// TIA Portal project "Blower_Speeds" (V19)
// Project for control of blower speed through variable frequency drive

(* hardware
DEVICE "S7-1200 station_1"  S7-1200 Station
   slot 0: "Rack_0"  S7-1200 Rack  Rack  V1.0
   slot 1: "PLC_1"  CPU 1212C AC/DC/Rly  6ES7 212-1BE40-0XB0  V4.6
DEVICE "HMI_1"  TP1200 Comfort
   slot 0: "HMI_1"  TP1200 Comfort  6AV2 124-0MC01-0AX0  17.0.0.0
   slot 1: "HMI_RT_1"  TP1200 Comfort  6AV2 124-0MC01-0AX0  17.0.0.0
   slot 5: "HMI_1.IE_CP_1"  PROFINET Interface  17.0.0.0
      slot 1: "PROFINET Interface_1"  PROFINET Interface
         slot 1: "Port_1"  Port
         slot 2: "Port_2"  Port
   slot 7: "HMI_1.MPI/DP_CP_1"  MPI/DP Interface  17.0.0.0
*)

// ===== PLC "PLC_1"  CPU 1212C AC/DC/Rly =====

VAR_GLOBAL   // PLC tag table "Inputs"
   "E_Stop" AT %I0.0 : Bool;   // Emergency stop
   "Start" AT %I0.2 : Bool;   // Pushbutton Start NO
   "Increase_Speed" AT %I0.4 : Bool;   // Pushbutton Increase NO
   "Decrease_Speed" AT %I0.3 : Bool;   // Pushbutton Decrease NO
   "Stop" AT %I0.1 : Bool;   // Pushbutton Stop NC
   "Tag_1" AT %M0.0 : Bool;
   "Tag_2" AT %M0.1 : Bool;
END_VAR

VAR_GLOBAL   // PLC tag table "Outputs"
   "Speed_1" AT %Q0.0 : Bool;   // Select Speed 1
   "Speed_2" AT %Q0.1 : Bool;   // Select Speed 2
   "Speed_3" AT %Q0.2 : Bool;   // Select Speed 3
   "Speed_4" AT %Q0.3 : Bool;   // Select Speed 4
END_VAR

// folder: DB

DATA_BLOCK "Data"   // DB1
TITLE = Data for Set Memories
{ S7_Optimized_Access := 'TRUE' }
AUTHOR : Stiven Perez
VERSION : 0.1
// Data for Set Memories
   VAR
      Start_Stop : Bool;   // Set-Reset Start or Stop Process
      P_Inc : Bool;
      N_Dec : Bool;
      QTime_1 : Bool;
      QTime_2 : Bool;
      QTime_3 : Bool;
      QTime_4 : Bool;
      CV_Speed : Int;
      Reset_Counter : Bool;
   END_VAR
BEGIN
END_DATA_BLOCK

DATA_BLOCK "Start_Stop_DB"   // DB2
{ S7_Optimized_Access := 'TRUE' }
VERSION : 0.1
// stored: InstanceOfName Start_Stop
"Start_Stop"
BEGIN
END_DATA_BLOCK

DATA_BLOCK "Inc_Dec_Speed_DB"   // DB3
{ S7_Optimized_Access := 'TRUE' }
AUTHOR : Stiven Perez
VERSION : 0.1
// stored: InstanceOfName Inc_Dec_Speed
"Inc_Dec_Speed"
BEGIN
END_DATA_BLOCK

DATA_BLOCK "Variables_HMI"   // DB4
TITLE = Variables for HMI
{ S7_Optimized_Access := 'TRUE' }
AUTHOR : Stiven Perez
VERSION : 0.1
   VAR
      Start_HMI : Bool;   // Start button HMI
      Stop_HMI : Bool;   // Stop button HMI
      Increase_HMI : Bool;   // Increase button HMI
      Decrease_HMI : Bool;   // Decrease button HMI
      Speed_1_HMI : Bool;   // Speed one
      Speed_2_HMI : Bool;   // Speed two
      Speed_3_HMI : Bool;   // Speed Three
      Speed_4_HMI : Bool;   // Speed four
   END_VAR
BEGIN
END_DATA_BLOCK

// folder: System blocks/Program resources

DATA_BLOCK "Timer_Speed1"   // DB6
{ S7_Optimized_Access := 'TRUE' }
AUTHOR : Simatic
FAMILY : IEC
NAME : IEC_TMR
VERSION : 1.0
// stored: InstanceOfName IEC_TIMER
"IEC_TIMER"
BEGIN
END_DATA_BLOCK

DATA_BLOCK "Timer_Speed2"   // DB7
{ S7_Optimized_Access := 'TRUE' }
AUTHOR : Simatic
FAMILY : IEC
NAME : IEC_TMR
VERSION : 1.0
// stored: InstanceOfName IEC_TIMER
"IEC_TIMER"
BEGIN
END_DATA_BLOCK

DATA_BLOCK "Timer_Speed3"   // DB8
{ S7_Optimized_Access := 'TRUE' }
AUTHOR : Simatic
FAMILY : IEC
NAME : IEC_TMR
VERSION : 1.0
// stored: InstanceOfName IEC_TIMER
"IEC_TIMER"
BEGIN
END_DATA_BLOCK

DATA_BLOCK "Timer_Speed4"   // DB9
{ S7_Optimized_Access := 'TRUE' }
AUTHOR : Simatic
FAMILY : IEC
NAME : IEC_TMR
VERSION : 1.0
// stored: InstanceOfName IEC_TIMER
"IEC_TIMER"
BEGIN
END_DATA_BLOCK

DATA_BLOCK "Counter_Speed"   // DB11
{ S7_Optimized_Access := 'TRUE' }
AUTHOR : Simatic
FAMILY : IEC
NAME : CNTR
VERSION : 1.0
// stored: InstanceOfName IEC_COUNTER
"IEC_COUNTER"
BEGIN
END_DATA_BLOCK

// folder: (top level)

ORGANIZATION_BLOCK "Main"   // OB1, LAD, ProgramCycle
TITLE = "Main Program Sweep (Cycle)"
{ S7_Optimized_Access := 'TRUE' }
VERSION : 0.1
   VAR_INPUT
      Initial_Call : Bool;   // Initial call of this OB
      Remanence : Bool;   // =True, if remanent data are available
   END_VAR
BEGIN

REGION Network 1: Start stop block
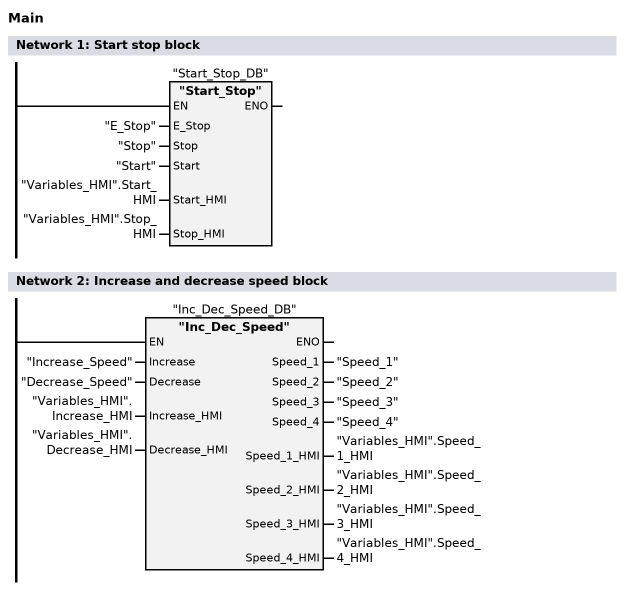
   RUNG wire#powerrail
      "Start_Stop_DB"(E_Stop := "E_Stop", Stop := "Stop", Start := "Start", Start_HMI := "Variables_HMI".Start_HMI, Stop_HMI := "Variables_HMI".Stop_HMI)
   END_RUNG
   // the same network as SCL:
   "Start_Stop_DB"(E_Stop := "E_Stop",   // "Start_Stop"
                   Stop := "Stop",
                   Start := "Start",
                   Start_HMI := "Variables_HMI".Start_HMI,
                   Stop_HMI := "Variables_HMI".Stop_HMI);
END_REGION

REGION Network 2: Increase and decrease speed block
   RUNG wire#powerrail
      "Inc_Dec_Speed_DB"(Increase := "Increase_Speed", Decrease := "Decrease_Speed", Increase_HMI := "Variables_HMI".Increase_HMI, Decrease_HMI := "Variables_HMI".Decrease_HMI, Speed_1 => "Speed_1", Speed_2 => "Speed_2", Speed_3 => "Speed_3", Speed_4 => "Speed_4", Speed_1_HMI => "Variables_HMI".Speed_1_HMI, Speed_2_HMI => "Variables_HMI".Speed_2_HMI, Speed_3_HMI => "Variables_HMI".Speed_3_HMI, Speed_4_HMI => "Variables_HMI".Speed_4_HMI)
   END_RUNG
   // the same network as SCL:
   "Inc_Dec_Speed_DB"(Increase := "Increase_Speed",   // "Inc_Dec_Speed"
                      Decrease := "Decrease_Speed",
                      Increase_HMI := "Variables_HMI".Increase_HMI,
                      Decrease_HMI := "Variables_HMI".Decrease_HMI,
                      Speed_1 => "Speed_1",
                      Speed_2 => "Speed_2",
                      Speed_3 => "Speed_3",
                      Speed_4 => "Speed_4",
                      Speed_1_HMI => "Variables_HMI".Speed_1_HMI,
                      Speed_2_HMI => "Variables_HMI".Speed_2_HMI,
                      Speed_3_HMI => "Variables_HMI".Speed_3_HMI,
                      Speed_4_HMI => "Variables_HMI".Speed_4_HMI);
END_REGION
END_ORGANIZATION_BLOCK

// folder: FB

FUNCTION_BLOCK "Inc_Dec_Speed"   // FB1, LAD
TITLE = Conditions to Increase and Decrease Speed
{ S7_Optimized_Access := 'TRUE' }
AUTHOR : Stiven Perez
VERSION : 0.1
// Conditions to select the respective speed
   VAR_INPUT
      Increase : Bool;
      Decrease : Bool;
      Increase_HMI : Bool;
      Decrease_HMI : Bool;
   END_VAR
   VAR_OUTPUT
      Speed_1 : Bool;
      Speed_2 : Bool;
      Speed_3 : Bool;
      Speed_4 : Bool;
      Speed_1_HMI : Bool;
      Speed_2_HMI : Bool;
      Speed_3_HMI : Bool;
      Speed_4_HMI : Bool;
   END_VAR
   VAR_TEMP   // added for the SCL form of the ladder/FBD networks
      _w1 : Bool;
      _w2 : Bool;
      _w3 : Bool;
      _w4 : Bool;
   END_VAR
BEGIN

REGION Network 1: Increase Speed
   // Conditions to increase or decrease speed
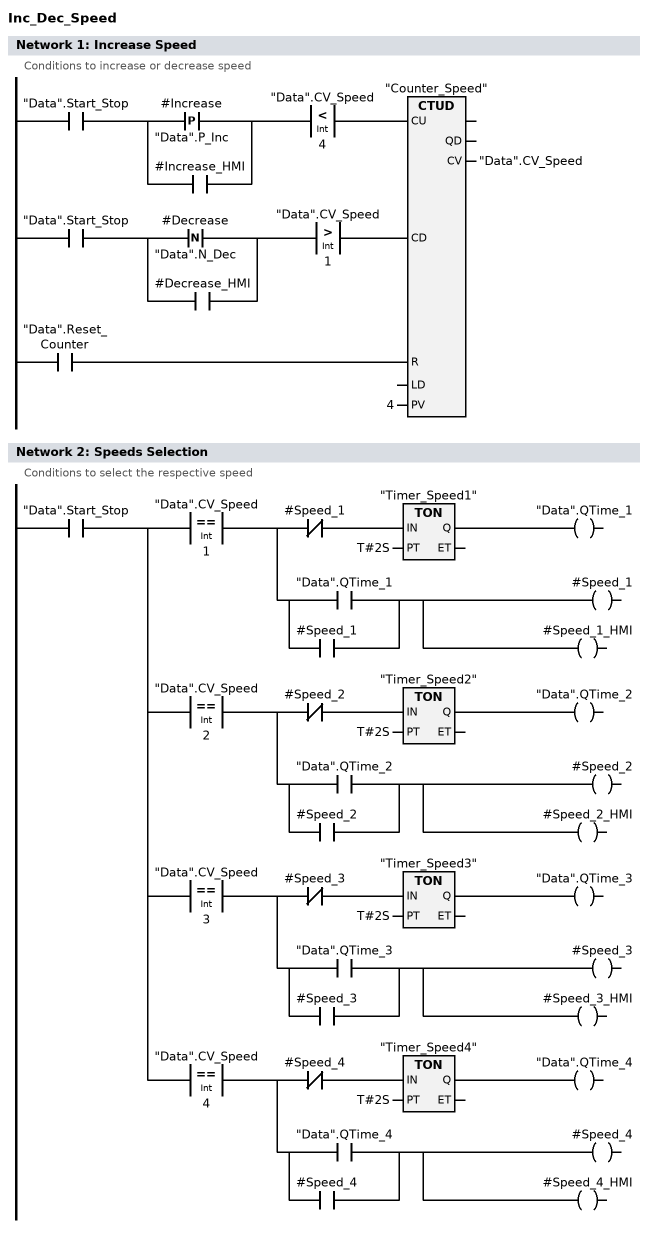
   #_w1 := "Data".Start_Stop AND #Increase AND NOT "Data".P_Inc;   // rising edge of #Increase
   "Data".P_Inc := #Increase;
   #_w2 := "Data".Start_Stop AND NOT #Decrease AND "Data".N_Dec;   // falling edge of #Decrease
   "Data".N_Dec := #Decrease;
   "Counter_Speed".CTUD(CU := (#_w1 OR ("Data".Start_Stop AND #Increase_HMI)) AND ("Data".CV_Speed < 4),
                        CD := (#_w2 OR ("Data".Start_Stop AND #Decrease_HMI)) AND ("Data".CV_Speed > 1),
                        R := "Data".Reset_Counter,
                        PV := 4,
                        CV => "Data".CV_Speed);
END_REGION

REGION Network 2: Speeds Selection
   // Conditions to select the respective speed
   #_w1 := "Data".Start_Stop AND ("Data".CV_Speed = 1);
   "Timer_Speed1".TON(IN := #_w1 AND NOT #Speed_1, PT := T#2S);
   "Data".QTime_1 := "Timer_Speed1".Q;
   #Speed_1 := #_w1 AND ("Data".QTime_1 OR #Speed_1);
   #Speed_1_HMI := #Speed_1;
   #_w2 := "Data".Start_Stop AND ("Data".CV_Speed = 2);
   "Timer_Speed2".TON(IN := #_w2 AND NOT #Speed_2, PT := T#2S);
   "Data".QTime_2 := "Timer_Speed2".Q;
   #Speed_2 := #_w2 AND ("Data".QTime_2 OR #Speed_2);
   #Speed_2_HMI := #Speed_2;
   #_w3 := "Data".Start_Stop AND ("Data".CV_Speed = 3);
   "Timer_Speed3".TON(IN := #_w3 AND NOT #Speed_3, PT := T#2S);
   "Data".QTime_3 := "Timer_Speed3".Q;
   #Speed_3 := #_w3 AND ("Data".QTime_3 OR #Speed_3);
   #Speed_3_HMI := #Speed_3;
   #_w4 := "Data".Start_Stop AND ("Data".CV_Speed = 4);
   "Timer_Speed4".TON(IN := #_w4 AND NOT #Speed_4, PT := T#2S);
   "Data".QTime_4 := "Timer_Speed4".Q;
   #Speed_4 := #_w4 AND ("Data".QTime_4 OR #Speed_4);
   #Speed_4_HMI := #Speed_4;
END_REGION
END_FUNCTION_BLOCK

FUNCTION_BLOCK "Start_Stop"   // FB2, LAD
TITLE = Start_Stop_Program
{ S7_Optimized_Access := 'TRUE' }
VERSION : 0.1
// Conditions to Start or stop all process
   VAR_INPUT
      E_Stop : Bool;
      Stop : Bool;
      Start : Bool;
      Start_HMI : Bool;
      Stop_HMI : Bool;
   END_VAR
   VAR_TEMP   // added for the SCL form of the ladder/FBD networks
      _w1 : Bool;
   END_VAR
BEGIN

REGION Network 1: Start Process
   // Start program
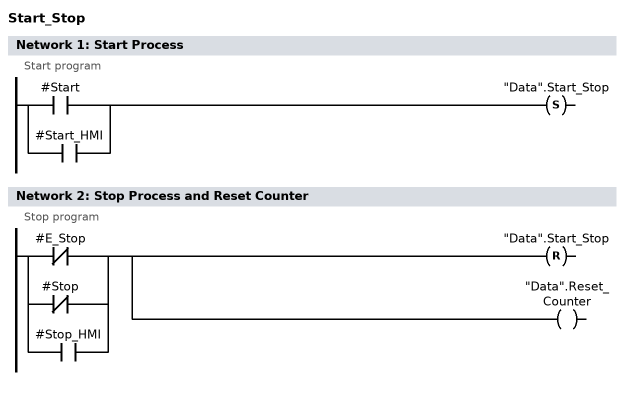
   RUNG wire#powerrail
      Contact( #Start )
      wire#w1
      S_Coil( "Data".Start_Stop )
   END_RUNG
   RUNG wire#powerrail
      Contact( #Start_HMI )
   END_RUNG wire#w1
   // the same network as SCL:
   IF #Start OR #Start_HMI THEN "Data".Start_Stop := TRUE; END_IF;
END_REGION

REGION Network 2: Stop Process and Reset Counter
   // Stop program
   RUNG wire#powerrail
      I_Contact( #E_Stop )
      wire#w1
      R_Coil( "Data".Start_Stop )
   END_RUNG
   RUNG wire#powerrail
      I_Contact( #Stop )
   END_RUNG wire#w1
   RUNG wire#powerrail
      Contact( #Stop_HMI )
   END_RUNG wire#w1
   RUNG wire#w1
      Coil( "Data".Reset_Counter )
   END_RUNG
   // the same network as SCL:
   #_w1 := NOT #E_Stop OR NOT #Stop OR #Stop_HMI;
   IF #_w1 THEN "Data".Start_Stop := FALSE; END_IF;
   "Data".Reset_Counter := #_w1;
END_REGION
END_FUNCTION_BLOCK

(* ===== HMI "HMI_RT_1" =====
system functions are stored by id; their names below are inferred from use
connection "HMI_Connection_1": ETHERNET, S7_1200_OMS

HMI tags "DATA_HMI"
   "Start" : Bool = PLC Variables_HMI.Start_HMI AT %DB1.DBW0, 100 ms
   "Stop" : Bool = PLC Variables_HMI.Stop_HMI AT %DB1.DBW0, 1 s
   "Increase" : Bool = PLC Variables_HMI.Increase_HMI AT %DB1.DBW0, 1 s
   "Decrease" : Bool = PLC Variables_HMI.Decrease_HMI AT %DB1.DBW0, 1 s
   "Speed_1" : Bool = PLC Variables_HMI.Speed_1_HMI AT %DB1.DBX0.0, 1 s
   "Speed_2" : Bool = PLC Variables_HMI.Speed_2_HMI AT %DB1.DBX0.0, 1 s
   "Speed_3" : Bool = PLC Variables_HMI.Speed_3_HMI AT %DB1.DBX0.0, 1 s
   "Speed_4" : Bool = PLC Variables_HMI.Speed_4_HMI AT %DB1.DBX0.0, 1 s
   "Set_Start" : Bool = PLC Data.Start_Stop AT %DB1.DBX0.0, 1 s

screen "Root screen" 1280x740, template "Template_1"
   on GenerateScreen: SetTag("Start", 1)
   TextField "Text field_1" at 484,43 size 320x37; Text 'Blower Speed Control'
   GraphicView "Graphic view_2" at 513,362 size 229x215; Picture "Graphic_2"
   GraphicView "Graphic view_6" at 132,192 size 119x126; Picture "Graphic_6"
      Visibility <- "Speed_1"
   GraphicView "Graphic view_1" at 432,191 size 119x126; Picture "Graphic_6"
      Visibility <- "Speed_2"
   GraphicView "Graphic view_3" at 767,191 size 119x126; Picture "Graphic_6"
      Visibility <- "Speed_3"
   GraphicView "Graphic view_4" at 1062,190 size 119x126; Picture "Graphic_6"
      Visibility <- "Speed_4"
   TextField "Text field_2" at 144,129 size 86x60; Text 'SPEED ONE'
      Appearance <- "Speed_1"
   TextField "Text field_3" at 452,129 size 86x60; Text 'SPEED TWO'
      Appearance <- "Speed_2"
   TextField "Text field_4" at 780,125 size 87x60; Text 'SPEED THREE'
      Appearance <- "Speed_3"
   TextField "Text field_5" at 1074,124 size 86x60; Text 'SPEED FOUR'
      Appearance <- "Speed_4"
   Button "Button_1" at 987,363 size 188x56; TextOff 'Increase Speed'
      on Press: function_b14e0dd5("Increase", 0)
   Button "Button_2" at 987,490 size 188x56; TextOff 'Decrease Speed'
      on Press: function_b14e0dd5("Decrease", 0)
   Button "Button_3" at 124,362 size 188x56; TextOff 'Start'
      on Press: SetBit("Start")
      on Release: ResetBit("Start")
      Appearance <- "Set_Start"
   Button "Button_4" at 125,490 size 188x56; TextOff 'Stop'
      on Press: SetBit("Stop")
      on Release: ResetBit("Stop")
      Appearance <- "Set_Start"
   GraphicView "Graphic view_7" at 130,193 size 120x127; Picture "Graphic_9"
      Visibility <- "Speed_1"
   GraphicView "Graphic view_5" at 430,192 size 120x127; Picture "Graphic_9"
      Visibility <- "Speed_2"
   GraphicView "Graphic view_8" at 764,192 size 120x127; Picture "Graphic_9"
      Visibility <- "Speed_3"
   GraphicView "Graphic view_9" at 1060,191 size 120x127; Picture "Graphic_9"
      Visibility <- "Speed_4"

Template "Template_1" 1280x740
   Button "Exit" at 1200,679 size 78x59; TextOff 'Exit'; PictureOff "ExitRuntime_TP1200_Comfort_TR"; PictureOn "ExitRuntime_TP1200_Comfort_TR"
      on Release: StopRuntime(0)
   Button "Template_Button" at 1120,679 size 78x59; TextOff 'Text'
   Button "Template_Button_1" at 1040,679 size 78x59; TextOff 'Text'
   Button "Template_Button_2" at 960,679 size 78x59; TextOff 'Text'
   Button "Template_Button_3" at 880,679 size 78x59; TextOff 'Text'
   Button "Template_Button_4" at 800,679 size 78x59; TextOff 'Text'
   Button "Template_Button_5" at 720,679 size 78x59; TextOff 'Text'
   Button "Template_Button_6" at 640,679 size 78x59; TextOff 'Text'
   Button "Template_Button_7" at 561,679 size 78x59; TextOff 'Text'
   Button "Template_Button_8" at 481,679 size 78x59; TextOff 'Text'
   Button "Template_Button_9" at 401,679 size 78x59; TextOff 'Text'
   Button "Template_Button_10" at 321,679 size 78x59; TextOff 'Text'
   Button "Template_Button_11" at 241,679 size 78x59; TextOff 'Text'
   Button "Template_Button_12" at 161,679 size 78x59; TextOff 'Text'
   Button "Alarms" at 81,679 size 78x59; TextOff 'Alarms'; PictureOff "AlarmDisplay_TP1200_Comfort_TR"; PictureOn "AlarmDisplay_TP1200_Comfort_TR"
      on Release: function_ef3f5d25("Alarm window_Unacknowledged", -1)
   Button "Start screen" at 1,679 size 78x59; TextOff 'Start screen'; PictureOff "NavigateHome_TP1200_Comfort_TR"; PictureOn "NavigateHome_TP1200_Comfort_TR"
      on Release: ActivateScreen("Root screen", 0)
*)